            ER_774 : Bool;   // Störung Hubantrieb FU 2: Reserve
            ER_775 : Bool;   // Störung Hubantrieb FU 2: Reserve
            ER_776_ : Bool;   // Störung Hubantrieb FU 2: Reserve
            ER_777 : Bool;   // Störung Hubantrieb FU 2: Reserve
            ER_778 : Bool;   // Störung Hubantrieb FU 2: Reserve
            ER_779 : Bool;   // Störung Hubantrieb FU 2: Reserve
            ER_780 : Bool;   // Störung Hubantrieb FU 2: Reserve
         END_STRUCT;
         Reserve_1 : Struct
            ER_401 : Bool;   // Reserve
            ER_402 : Bool;   // Reserve
            ER_403 : Bool;   // Reserve
            ER_404 : Bool;   // Reserve
            ER_405 : Bool;   // Reserve
            ER_406 : Bool;   // Reserve
            ER_407 : Bool;   // Reserve
            ER_408 : Bool;   // Reserve
            ER_409 : Bool;   // Reserve
            ER_410 : Bool;   // Reserve
            ER_411 : Bool;   // Reserve
            ER_412 : Bool;   // Reserve
            ER_413 : Bool;   // Reserve
            ER_414 : Bool;   // Reserve
            ER_415 : Bool;   // Reserve
            ER_416 : Bool;   // Reserve
         END_STRUCT;
         Reserve_2 : Struct
            ER_417 : Bool;   // Reserve
            ER_418 : Bool;   // Reserve
            ER_419 : Bool;   // Reserve
            ER_420 : Bool;   // Reserve
            ER_421 : Bool;   // Reserve
            ER_422 : Bool;   // Reserve
            ER_423 : Bool;   // Reserve
            ER_424 : Bool;   // Reserve
            ER_425 : Bool;   // Reserve
            ER_426 : Bool;   // Reserve
            ER_427 : Bool;   // Reserve
            ER_428 : Bool;   // Reserve
            ER_429 : Bool;   // Reserve
            ER_430 : Bool;   // Reserve
            ER_431 : Bool;   // Reserve
            ER_432 : Bool;   // Reserve
         END_STRUCT;
         Reserve_3 : Struct
            ER_433 : Bool;   // Reserve
            ER_434 : Bool;   // Reserve
            ER_435 : Bool;   // Reserve
            ER_436 : Bool;   // Reserve
            ER_437 : Bool;   // Reserve
            ER_438 : Bool;   // Reserve
            ER_439 : Bool;   // Reserve
            ER_440 : Bool;   // Reserve
            ER_441 : Bool;   // Reserve
            ER_442 : Bool;   // Reserve
            ER_443 : Bool;   // Reserve
            ER_444 : Bool;   // Reserve
            ER_445 : Bool;   // Reserve
            ER_446 : Bool;   // Reserve
            ER_447 : Bool;   // Reserve
            ER_448 : Bool;   // Reserve
         END_STRUCT;
         Reserve_4 : Struct
            ER_449 : Bool;   // Reserve
            ER_450 : Bool;   // Reserve
            ER_451 : Bool;   // Reserve
            ER_452 : Bool;   // Reserve
            ER_453 : Bool;   // Reserve
            ER_454 : Bool;   // Reserve
            ER_455 : Bool;   // Reserve
            ER_456 : Bool;   // Reserve
            ER_457 : Bool;   // Reserve
            ER_458 : Bool;   // Reserve
            ER_459 : Bool;   // Reserve
            ER_460 : Bool;   // Reserve
            ER_461 : Bool;   // Reserve
            ER_462 : Bool;   // Reserve
            ER_463 : Bool;   // Reserve
            ER_464 : Bool;   // Reserve
         END_STRUCT;
         Reserve_5 : Struct
            ER_465 : Bool;   // Reserve
            ER_466 : Bool;   // Reserve
            ER_467 : Bool;   // Reserve
            ER_468 : Bool;   // Reserve
            ER_469 : Bool;   // Reserve
            ER_470 : Bool;   // Reserve
            ER_471 : Bool;   // Reserve
            ER_472 : Bool;   // Reserve
            ER_473 : Bool;   // Reserve
            ER_474 : Bool;   // Reserve
            ER_475 : Bool;   // Reserve
            ER_476 : Bool;   // Reserve
            ER_477 : Bool;   // Reserve
            ER_478 : Bool;   // Reserve
            ER_479 : Bool;   // Reserve
            ER_480 : Bool;   // Reserve
         END_STRUCT;
         Reserve_6 : Struct   // Meldungen Reserve
            ER_301 : Bool;   // Reserve
            ER_302 : Bool;   // Reserve
            ER_303 : Bool;   // Reserve
            ER_304 : Bool;   // Reserve
            ER_305 : Bool;   // Reserve
            ER_306 : Bool;   // Reserve
            ER_307 : Bool;   // Reserve
            ER_308 : Bool;   // Reserve
            ER_309 : Bool;   // Reserve
            ER_310 : Bool;   // Reserve
            ER_311 : Bool;   // Reserve
            ER_312 : Bool;   // Reserve
            ER_313 : Bool;   // Reserve
            ER_314 : Bool;   // Reserve
            ER_315 : Bool;   // Reserve
            ER_316 : Bool;   // Reserve
         END_STRUCT;
         Reserve_7 : Struct   // Meldungen Reserve
            ER_317 : Bool;   // Reserve
            ER_318 : Bool;   // Reserve
            ER_319 : Bool;   // Reserve
            ER_320 : Bool;   // Reserve
            ER_321 : Bool;   // Reserve
            ER_322 : Bool;   // Reserve
            ER_323 : Bool;   // Reserve
            ER_324 : Bool;   // Reserve
            ER_325 : Bool;   // Reserve
            ER_326 : Bool;   // Reserve
            ER_327 : Bool;   // Reserve
            ER_328 : Bool;   // Reserve
            ER_329 : Bool;   // Reserve
            ER_330 : Bool;   // Reserve
            ER_331 : Bool;   // Reserve
            ER_332 : Bool;   // Reserve
         END_STRUCT;
         Reserve_8 : Struct   // FU Reserve
            ER_333 : Bool;   // Störung Reserve FU 1: Überstrom
            ER_334 : Bool;   // Störung Reserve FU 1: Zwischenkreisspannung Überspannung
            ER_335 : Bool;   // Störung Reserve FU 1: Zwischenkreisspannung Unterspannung
            ER_336 : Bool;   // Störung Reserve FU 1: Übertemperatur Kühlkörper Wechselrichter
            ER_337 : Bool;   // Störung Reserve FU 1: Motordatenidentifikation fehlerhaft
            ER_338 : Bool;   // Störung Reserve FU 1: Erdschluss
            ER_339 : Bool;   // Störung Reserve FU 1: Reserve
            ER_340 : Bool;   // Störung Reserve FU 1: Führung durch PLC fehlt
            ER_341 : Bool;   // Störung Reserve FU 1: Reserve
            ER_342 : Bool;   // Störung Reserve FU 1: Reserve
            ER_343 : Bool;   // Störung Reserve FU 1: Reserve
            ER_344_ : Bool;   // Störung Reserve FU 1: Reserve
            ER_345 : Bool;   // Störung Reserve FU 1: Reserve
            ER_346 : Bool;   // Störung Reserve FU 1: Reserve
            ER_347 : Bool;   // Störung Reserve FU 1: Reserve
            ER_348 : Bool;   // Störung Reserve FU 1: Reserve
         END_STRUCT;
         Reserve_9 : Struct
            ER_349 : Bool;   // Reserve
            ER_350 : Bool;   // Reserve
            ER_351 : Bool;   // Reserve
            ER_352 : Bool;   // Reserve
            ER_353 : Bool;   // Reserve
            ER_354 : Bool;   // Reserve
            ER_355 : Bool;   // Reserve
            ER_356 : Bool;   // Reserve
            ER_357 : Bool;   // Reserve
            ER_358 : Bool;   // Reserve
            ER_359 : Bool;   // Reserve
            ER_360 : Bool;   // Reserve
            ER_361 : Bool;   // Reserve
            ER_362 : Bool;   // Reserve
            ER_363 : Bool;   // Reserve
            ER_364 : Bool;   // Reserve
         END_STRUCT;
         Reserve_10 : Struct   // FU Reserve
            ER_365 : Bool;   // Störung Reserve FU 2: Überstrom
            ER_366 : Bool;   // Störung Reserve FU 2: Zwischenkreisspannung Überspannung
            ER_367 : Bool;   // Störung Reserve FU 2: Zwischenkreisspannung Unterspannung
            ER_368 : Bool;   // Störung Reserve FU 2: Übertemperatur Kühlkörper Wechselrichter
            ER_369 : Bool;   // Störung Reserve FU 2: Motordatenidentifikation fehlerhaft
            ER_370 : Bool;   // Störung Reserve FU 2: Erdschluss
            ER_371 : Bool;   // Störung Reserve FU 2: Reserve
            ER_372 : Bool;   // Störung Reserve FU 2: Führung durch PLC fehlt
            ER_373 : Bool;   // Störung Reserve FU 2: Reserve
            ER_374 : Bool;   // Störung Reserve FU 2: Reserve
            ER_375 : Bool;   // Störung Reserve FU 2: Reserve
            ER_376 : Bool;   // Störung Reserve FU 2: Reserve
            ER_377 : Bool;   // Störung Reserve FU 2: Reserve
            ER_378 : Bool;   // Störung Reserve FU 2: Reserve
            ER_379 : Bool;   // Störung Reserve FU 2: Reserve
            ER_380 : Bool;   // Störung Reserve FU 2: Reserve
         END_STRUCT;
         SDC : Struct   // SDC Störungs
            ER_901 : Bool;   // Reserve
            ER_902 : Bool;   // Reserve
            ER_903 : Bool;   // Störung SDC Positionssprung
            ER_904 : Bool;   // Störung SDC keine Sektion gefunden
            ER_905 : Bool;   // Störung SDC Kommandos nicht plausibel
            ER_906 : Bool;   // Störung SDC Positionsgrenzen
            ER_907 : Bool;   // Störung SDC falsche EMS Nummer
            ER_908 : Bool;   // Störung SDC falsche Sektion Nummer
            ER_909 : Bool;   // Reserve
            ER_910 : Bool;   // Reserve
            ER_911 : Bool;   // Reserve
            ER_912 : Bool;   // Reserve
            ER_913 : Bool;   // Reserve
            ER_914 : Bool;   // Reserve
            ER_915 : Bool;   // Reserve
            ER_916 : Bool;   // Reserve
         END_STRUCT;
      END_STRUCT;
      EMS_ER_WORDs : Array[1..200] of Struct   // EMS Störung WORDs
         ER_WORD : Array[0..24] of Word;   // Störworte
      END_STRUCT;
      SDC : Struct
         ER_917 : Bool;   // Störung SDC Kommunikation mit Anlagensteuerung
         ER_918 : Bool;   // Störung SDC Safety Kommunikation mit Anlagensteuerung
         ER_919 : Bool;   // Störung SDC Reserve
         ER_920 : Bool;   // Störung SDC Reserve
         ER_921 : Bool;   // Störung SDC Reserve
         ER_922 : Bool;   // Störung SDC Reserve
         ER_923 : Bool;   // Störung SDC Reserve
         ER_924 : Bool;   // Störung SDC Reserve
         ER_925 : Bool;   // Störung SDC OB80 Zykluszeit
         ER_926 : Bool;   // Störung SDC OB82 Diagnosealarm
         ER_927 : Bool;   // Störung SDC OB83 Baugruppenwechsel
         ER_928 : Bool;   // Störung SDC OB86 Baugruppenträger ausgefallen
         ER_929 : Bool;   // Störung SDC OB121 Programmierfehler
         ER_930 : Bool;   // Störung SDC OB122 Peripherie-Zugriff
         ER_931 : Bool;   // Störung SDC Reserve
         ER_932 : Bool;   // Störung SDC Reserve
      END_STRUCT;
   END_VAR
BEGIN
END_DATA_BLOCK

DATA_BLOCK "DB_SDC_ERRORS_STAT"   // DB3724
{ S7_Optimized_Access := 'FALSE' }
VERSION : 0.1
   VAR
      HEADER : Struct   // Struktur für Datenheader // nicht verschieben
         DB_NR : Int := 3724;   // DB Nummer
         MIN_NR_FAULT_STAT : Int := 1;   // Niedrigste Fehler Nummer im Daten DB
         MAX_NR_FAULT_STAT : Int := 200;   // Höchste Fehler Nummer im Daten DB
         START_FAULT_STAT : Int := 20;   // Startadresse der Fehler Daten im Daten DB
         LAENGE_FAULT_STAT : Int := 28;   // Länge Fehler Daten
         FAULT_PRO_SEITE_HMI : Int := 10;   // Reserve
         RES12 : Int := 0;   // Reserve
         RES14 : Int := 0;   // Reserve
         RES16 : Int := 0;   // Reserve
         LOAD : Bool := FALSE;   // "0" zum laden des DB auf CPU
         RESET_ARCH : Bool := FALSE;   // Archiv löschen
      END_STRUCT;
      ER_ARCHIV : Array[1..1000] of "UDT_SDC_ERROR_STAT";   // Error Archiv
      ER_AKT : Array[1..200] of Struct   // Error aktiv EMS
         ER_TRIGER : Word;   // Error auslösen Aktiv von EMS
         ER_STAT : Array[1..4] of "UDT_SDC_TS_IF_STATUS_VAL";   // Error Status Aktiv EMS
      END_STRUCT;
   END_VAR
BEGIN
   ER_ARCHIV[1].EMS_TS_STAT_VAL.EMS_ID := 0;
   ER_ARCHIV[1].EMS_TS_STAT_VAL.PROFIL := 0;
   ER_ARCHIV[1].EMS_TS_STAT_VAL.DRIVE_POS := 0;
   ER_ARCHIV[1].EMS_TS_STAT_VAL.HOIST_POS := 0;
   ER_ARCHIV[1].EMS_TS_STAT_VAL.ERROR := 0;
   ER_ARCHIV[1].EMS_TS_STAT_VAL.DRIVE_POS_PERC := 0;
   ER_ARCHIV[1].EMS_TS_STAT_VAL.SEK := 0;
   ER_ARCHIV[1].ER._901_ER_SUM := FALSE;
   ER_ARCHIV[1].ER._902_ER_SUM_SDC := FALSE;
   ER_ARCHIV[1].ER._903_ER_BC_JUMP := FALSE;
   ER_ARCHIV[1].ER._904_ER_NO_SEK := FALSE;
   ER_ARCHIV[1].ER._905_ER_COMMAND := FALSE;
   ER_ARCHIV[1].ER._906_ER_BC_LIM := FALSE;
   ER_ARCHIV[1].ER._907_ER_EMS_ID := FALSE;
   ER_ARCHIV[1].ER._908_ER_SEK_NR := FALSE;
   ER_ARCHIV[1].ER._909_ER_LIFE := FALSE;
   ER_ARCHIV[1].ER._910_ER_BUS := FALSE;
   ER_ARCHIV[1].ER._911 := FALSE;
   ER_ARCHIV[1].ER._912 := FALSE;
   ER_ARCHIV[1].ER._913 := FALSE;
   ER_ARCHIV[1].ER._914 := FALSE;
   ER_ARCHIV[1].ER._915 := FALSE;
   ER_ARCHIV[1].ER._916 := FALSE;
   ER_ARCHIV[1].Spare := 0;
   ER_ARCHIV[1].ER_DATE := DT#1990-01-01-00:00:00;
   ER_ARCHIV[2].EMS_TS_STAT_VAL.EMS_ID := 0;
   ER_ARCHIV[2].EMS_TS_STAT_VAL.PROFIL := 0;
   ER_ARCHIV[2].EMS_TS_STAT_VAL.DRIVE_POS := 0;
   ER_ARCHIV[2].EMS_TS_STAT_VAL.HOIST_POS := 0;
   ER_ARCHIV[2].EMS_TS_STAT_VAL.ERROR := 0;
   ER_ARCHIV[2].EMS_TS_STAT_VAL.DRIVE_POS_PERC := 0;
   ER_ARCHIV[2].EMS_TS_STAT_VAL.SEK := 0;
   ER_ARCHIV[2].ER._901_ER_SUM := FALSE;
   ER_ARCHIV[2].ER._902_ER_SUM_SDC := FALSE;
   ER_ARCHIV[2].ER._903_ER_BC_JUMP := FALSE;
   ER_ARCHIV[2].ER._904_ER_NO_SEK := FALSE;
   ER_ARCHIV[2].ER._905_ER_COMMAND := FALSE;
   ER_ARCHIV[2].ER._906_ER_BC_LIM := FALSE;
   ER_ARCHIV[2].ER._907_ER_EMS_ID := FALSE;
   ER_ARCHIV[2].ER._908_ER_SEK_NR := FALSE;
   ER_ARCHIV[2].ER._909_ER_LIFE := FALSE;
   ER_ARCHIV[2].ER._910_ER_BUS := FALSE;
   ER_ARCHIV[2].ER._911 := FALSE;
   ER_ARCHIV[2].ER._912 := FALSE;
   ER_ARCHIV[2].ER._913 := FALSE;
   ER_ARCHIV[2].ER._914 := FALSE;
   ER_ARCHIV[2].ER._915 := FALSE;
   ER_ARCHIV[2].ER._916 := FALSE;
   ER_ARCHIV[2].Spare := 0;
   ER_ARCHIV[2].ER_DATE := DT#1990-01-01-00:00:00;
   ER_ARCHIV[3].EMS_TS_STAT_VAL.EMS_ID := 0;
   ER_ARCHIV[3].EMS_TS_STAT_VAL.PROFIL := 0;
   ER_ARCHIV[3].EMS_TS_STAT_VAL.DRIVE_POS := 0;
   ER_ARCHIV[3].EMS_TS_STAT_VAL.HOIST_POS := 0;
   ER_ARCHIV[3].EMS_TS_STAT_VAL.ERROR := 0;
   ER_ARCHIV[3].EMS_TS_STAT_VAL.DRIVE_POS_PERC := 0;
   ER_ARCHIV[3].EMS_TS_STAT_VAL.SEK := 0;
   ER_ARCHIV[3].ER._901_ER_SUM := FALSE;
   ER_ARCHIV[3].ER._902_ER_SUM_SDC := FALSE;
   ER_ARCHIV[3].ER._903_ER_BC_JUMP := FALSE;
   ER_ARCHIV[3].ER._904_ER_NO_SEK := FALSE;
   ER_ARCHIV[3].ER._905_ER_COMMAND := FALSE;
   ER_ARCHIV[3].ER._906_ER_BC_LIM := FALSE;
   ER_ARCHIV[3].ER._907_ER_EMS_ID := FALSE;
   ER_ARCHIV[3].ER._908_ER_SEK_NR := FALSE;
   ER_ARCHIV[3].ER._909_ER_LIFE := FALSE;
   ER_ARCHIV[3].ER._910_ER_BUS := FALSE;
   ER_ARCHIV[3].ER._911 := FALSE;
   ER_ARCHIV[3].ER._912 := FALSE;
   ER_ARCHIV[3].ER._913 := FALSE;
   ER_ARCHIV[3].ER._914 := FALSE;
   ER_ARCHIV[3].ER._915 := FALSE;
   ER_ARCHIV[3].ER._916 := FALSE;
   ER_ARCHIV[3].Spare := 0;
   ER_ARCHIV[3].ER_DATE := DT#1990-01-01-00:00:00;
   ER_ARCHIV[4].EMS_TS_STAT_VAL.EMS_ID := 0;
   ER_ARCHIV[4].EMS_TS_STAT_VAL.PROFIL := 0;
   ER_ARCHIV[4].EMS_TS_STAT_VAL.DRIVE_POS := 0;
   ER_ARCHIV[4].EMS_TS_STAT_VAL.HOIST_POS := 0;
   ER_ARCHIV[4].EMS_TS_STAT_VAL.ERROR := 0;
   ER_ARCHIV[4].EMS_TS_STAT_VAL.DRIVE_POS_PERC := 0;
   ER_ARCHIV[4].EMS_TS_STAT_VAL.SEK := 0;
   ER_ARCHIV[4].ER._901_ER_SUM := FALSE;
   ER_ARCHIV[4].ER._902_ER_SUM_SDC := FALSE;
   ER_ARCHIV[4].ER._903_ER_BC_JUMP := FALSE;
   ER_ARCHIV[4].ER._904_ER_NO_SEK := FALSE;
   ER_ARCHIV[4].ER._905_ER_COMMAND := FALSE;
   ER_ARCHIV[4].ER._906_ER_BC_LIM := FALSE;
   ER_ARCHIV[4].ER._907_ER_EMS_ID := FALSE;
   ER_ARCHIV[4].ER._908_ER_SEK_NR := FALSE;
   ER_ARCHIV[4].ER._909_ER_LIFE := FALSE;
   ER_ARCHIV[4].ER._910_ER_BUS := FALSE;
   ER_ARCHIV[4].ER._911 := FALSE;
   ER_ARCHIV[4].ER._912 := FALSE;
   ER_ARCHIV[4].ER._913 := FALSE;
   ER_ARCHIV[4].ER._914 := FALSE;
   ER_ARCHIV[4].ER._915 := FALSE;
   ER_ARCHIV[4].ER._916 := FALSE;
   ER_ARCHIV[4].Spare := 0;
   ER_ARCHIV[4].ER_DATE := DT#1990-01-01-00:00:00;
   ER_ARCHIV[5].EMS_TS_STAT_VAL.EMS_ID := 0;
   ER_ARCHIV[5].EMS_TS_STAT_VAL.PROFIL := 0;
   ER_ARCHIV[5].EMS_TS_STAT_VAL.DRIVE_POS := 0;
   ER_ARCHIV[5].EMS_TS_STAT_VAL.HOIST_POS := 0;
   ER_ARCHIV[5].EMS_TS_STAT_VAL.ERROR := 0;
   ER_ARCHIV[5].EMS_TS_STAT_VAL.DRIVE_POS_PERC := 0;
   ER_ARCHIV[5].EMS_TS_STAT_VAL.SEK := 0;
   ER_ARCHIV[5].ER._901_ER_SUM := FALSE;
   ER_ARCHIV[5].ER._902_ER_SUM_SDC := FALSE;
   ER_ARCHIV[5].ER._903_ER_BC_JUMP := FALSE;
   ER_ARCHIV[5].ER._904_ER_NO_SEK := FALSE;
   ER_ARCHIV[5].ER._905_ER_COMMAND := FALSE;
   ER_ARCHIV[5].ER._906_ER_BC_LIM := FALSE;
   ER_ARCHIV[5].ER._907_ER_EMS_ID := FALSE;
   ER_ARCHIV[5].ER._908_ER_SEK_NR := FALSE;
   ER_ARCHIV[5].ER._909_ER_LIFE := FALSE;
   ER_ARCHIV[5].ER._910_ER_BUS := FALSE;
   ER_ARCHIV[5].ER._911 := FALSE;
   ER_ARCHIV[5].ER._912 := FALSE;
   ER_ARCHIV[5].ER._913 := FALSE;
   ER_ARCHIV[5].ER._914 := FALSE;
   ER_ARCHIV[5].ER._915 := FALSE;
   ER_ARCHIV[5].ER._916 := FALSE;
   ER_ARCHIV[5].Spare := 0;
   ER_ARCHIV[5].ER_DATE := DT#1990-01-01-00:00:00;
   ER_ARCHIV[6].EMS_TS_STAT_VAL.EMS_ID := 0;
   ER_ARCHIV[6].EMS_TS_STAT_VAL.PROFIL := 0;
   ER_ARCHIV[6].EMS_TS_STAT_VAL.DRIVE_POS := 0;
   ER_ARCHIV[6].EMS_TS_STAT_VAL.HOIST_POS := 0;
   ER_ARCHIV[6].EMS_TS_STAT_VAL.ERROR := 0;
   ER_ARCHIV[6].EMS_TS_STAT_VAL.DRIVE_POS_PERC := 0;
   ER_ARCHIV[6].EMS_TS_STAT_VAL.SEK := 0;
   ER_ARCHIV[6].ER._901_ER_SUM := FALSE;
   ER_ARCHIV[6].ER._902_ER_SUM_SDC := FALSE;
   ER_ARCHIV[6].ER._903_ER_BC_JUMP := FALSE;
   ER_ARCHIV[6].ER._904_ER_NO_SEK := FALSE;
   ER_ARCHIV[6].ER._905_ER_COMMAND := FALSE;
   ER_ARCHIV[6].ER._906_ER_BC_LIM := FALSE;
   ER_ARCHIV[6].ER._907_ER_EMS_ID := FALSE;
   ER_ARCHIV[6].ER._908_ER_SEK_NR := FALSE;
   ER_ARCHIV[6].ER._909_ER_LIFE := FALSE;
   ER_ARCHIV[6].ER._910_ER_BUS := FALSE;
   ER_ARCHIV[6].ER._911 := FALSE;
   ER_ARCHIV[6].ER._912 := FALSE;
   ER_ARCHIV[6].ER._913 := FALSE;
   ER_ARCHIV[6].ER._914 := FALSE;
   ER_ARCHIV[6].ER._915 := FALSE;
   ER_ARCHIV[6].ER._916 := FALSE;
   ER_ARCHIV[6].Spare := 0;
   ER_ARCHIV[6].ER_DATE := DT#1990-01-01-00:00:00;
   ER_ARCHIV[7].EMS_TS_STAT_VAL.EMS_ID := 0;
   ER_ARCHIV[7].EMS_TS_STAT_VAL.PROFIL := 0;
   ER_ARCHIV[7].EMS_TS_STAT_VAL.DRIVE_POS := 0;
   ER_ARCHIV[7].EMS_TS_STAT_VAL.HOIST_POS := 0;
   ER_ARCHIV[7].EMS_TS_STAT_VAL.ERROR := 0;
   ER_ARCHIV[7].EMS_TS_STAT_VAL.DRIVE_POS_PERC := 0;
   ER_ARCHIV[7].EMS_TS_STAT_VAL.SEK := 0;
   ER_ARCHIV[7].ER._901_ER_SUM := FALSE;
   ER_ARCHIV[7].ER._902_ER_SUM_SDC := FALSE;
   ER_ARCHIV[7].ER._903_ER_BC_JUMP := FALSE;
   ER_ARCHIV[7].ER._904_ER_NO_SEK := FALSE;
   ER_ARCHIV[7].ER._905_ER_COMMAND := FALSE;
   ER_ARCHIV[7].ER._906_ER_BC_LIM := FALSE;
   ER_ARCHIV[7].ER._907_ER_EMS_ID := FALSE;
   ER_ARCHIV[7].ER._908_ER_SEK_NR := FALSE;
   ER_ARCHIV[7].ER._909_ER_LIFE := FALSE;
   ER_ARCHIV[7].ER._910_ER_BUS := FALSE;
   ER_ARCHIV[7].ER._911 := FALSE;
   ER_ARCHIV[7].ER._912 := FALSE;
   ER_ARCHIV[7].ER._913 := FALSE;
   ER_ARCHIV[7].ER._914 := FALSE;
   ER_ARCHIV[7].ER._915 := FALSE;
   ER_ARCHIV[7].ER._916 := FALSE;
   ER_ARCHIV[7].Spare := 0;
   ER_ARCHIV[7].ER_DATE := DT#1990-01-01-00:00:00;
   ER_ARCHIV[8].EMS_TS_STAT_VAL.EMS_ID := 0;
   ER_ARCHIV[8].EMS_TS_STAT_VAL.PROFIL := 0;
   ER_ARCHIV[8].EMS_TS_STAT_VAL.DRIVE_POS := 0;
   ER_ARCHIV[8].EMS_TS_STAT_VAL.HOIST_POS := 0;
   ER_ARCHIV[8].EMS_TS_STAT_VAL.ERROR := 0;
   ER_ARCHIV[8].EMS_TS_STAT_VAL.DRIVE_POS_PERC := 0;
   ER_ARCHIV[8].EMS_TS_STAT_VAL.SEK := 0;
   ER_ARCHIV[8].ER._901_ER_SUM := FALSE;
   ER_ARCHIV[8].ER._902_ER_SUM_SDC := FALSE;
   ER_ARCHIV[8].ER._903_ER_BC_JUMP := FALSE;
   ER_ARCHIV[8].ER._904_ER_NO_SEK := FALSE;
   ER_ARCHIV[8].ER._905_ER_COMMAND := FALSE;
   ER_ARCHIV[8].ER._906_ER_BC_LIM := FALSE;
   ER_ARCHIV[8].ER._907_ER_EMS_ID := FALSE;
   ER_ARCHIV[8].ER._908_ER_SEK_NR := FALSE;
   ER_ARCHIV[8].ER._909_ER_LIFE := FALSE;
   ER_ARCHIV[8].ER._910_ER_BUS := FALSE;
   ER_ARCHIV[8].ER._911 := FALSE;
   ER_ARCHIV[8].ER._912 := FALSE;
   ER_ARCHIV[8].ER._913 := FALSE;
   ER_ARCHIV[8].ER._914 := FALSE;
   ER_ARCHIV[8].ER._915 := FALSE;
   ER_ARCHIV[8].ER._916 := FALSE;
   ER_ARCHIV[8].Spare := 0;
   ER_ARCHIV[8].ER_DATE := DT#1990-01-01-00:00:00;
   // 30600 more start values not shown
END_DATA_BLOCK

DATA_BLOCK "DB_SDC_EMS_SIM"   // DB3726
{ S7_Optimized_Access := 'FALSE' }
VERSION : 0.1
   VAR
      HEADER : Struct   // Struktur für Datenheader // nicht verschieben
         DB_NR : Int := 3726;   // DB Nummer
         MIN_NR_EMS : Int := 1;   // Niedrigste EMS Nummer im Daten DB
         MAX_NR_EMS : Int := 200;   // Höchste EMS Nummer im Daten DB
         START_DAT : Int := 40;   // Startadresse der EMS Daten im Daten DB
         LAENGE_EMS : Int := 40;   // Länge Eingänge pro EMS
         RES10 : Int := 0;   // Reserve
         RES12 : Int := 0;   // Reserve
         RES14 : Int := 0;   // Reserve
         RES16 : Int := 0;   // Reserve
         RES18 : Int := 0;   // Reserve
      END_STRUCT;
      PAR : Struct   // Parameter Simulation
         BARCODE_START : DInt := 1;   // min Barcodevalue
         BARCODE_ENDE : DInt := 500000;   // max Barcodevalue
         HUB_START : Int := 0;   // min Hoistvalue
         HUB_ENDE : Int := 4010;   // max Hoistvalue
         LEAP_AKT : Array[1..20] of Bool;   // Leap Aktiv
         LEAP_HIGH_LOW : Array[1..20] of Bool;   // Leap Aktiv
         ON : Bool := TRUE;   // Simulation ON "1"
         RES18 : Int := 0;   // Reserve
      END_STRUCT;
      EMS : Array[1..200] of "UDT_EMS_IF_Q";   // EMS Simulation Eingänge
      EMS_TEMP : "UDT_EMS_IF_Q";
   END_VAR
BEGIN
   PAR.LEAP_AKT[1] := TRUE;
   PAR.LEAP_AKT[2] := TRUE;
   PAR.LEAP_AKT[3] := TRUE;
   PAR.LEAP_HIGH_LOW[1] := TRUE;
   PAR.LEAP_HIGH_LOW[2] := FALSE;
   PAR.LEAP_HIGH_LOW[3] := TRUE;
   PAR.LEAP_AKT[4] := FALSE;
   PAR.LEAP_AKT[5] := FALSE;
   PAR.LEAP_AKT[6] := FALSE;
   PAR.LEAP_AKT[7] := FALSE;
   PAR.LEAP_AKT[8] := FALSE;
   PAR.LEAP_AKT[9] := FALSE;
   PAR.LEAP_AKT[10] := FALSE;
   PAR.LEAP_AKT[11] := FALSE;
   PAR.LEAP_AKT[12] := FALSE;
   PAR.LEAP_AKT[13] := FALSE;
   PAR.LEAP_AKT[14] := FALSE;
   PAR.LEAP_AKT[15] := FALSE;
   PAR.LEAP_AKT[16] := FALSE;
   PAR.LEAP_AKT[17] := FALSE;
   PAR.LEAP_AKT[18] := FALSE;
   PAR.LEAP_AKT[19] := FALSE;
   PAR.LEAP_AKT[20] := FALSE;
   PAR.LEAP_HIGH_LOW[4] := FALSE;
   PAR.LEAP_HIGH_LOW[5] := FALSE;
   PAR.LEAP_HIGH_LOW[6] := FALSE;
   PAR.LEAP_HIGH_LOW[7] := FALSE;
   PAR.LEAP_HIGH_LOW[8] := FALSE;
   PAR.LEAP_HIGH_LOW[9] := FALSE;
   PAR.LEAP_HIGH_LOW[10] := FALSE;
   PAR.LEAP_HIGH_LOW[11] := FALSE;
   PAR.LEAP_HIGH_LOW[12] := FALSE;
   PAR.LEAP_HIGH_LOW[13] := FALSE;
   PAR.LEAP_HIGH_LOW[14] := FALSE;
   PAR.LEAP_HIGH_LOW[15] := FALSE;
   PAR.LEAP_HIGH_LOW[16] := FALSE;
   PAR.LEAP_HIGH_LOW[17] := FALSE;
   PAR.LEAP_HIGH_LOW[18] := FALSE;
   PAR.LEAP_HIGH_LOW[19] := FALSE;
   PAR.LEAP_HIGH_LOW[20] := FALSE;
   EMS[1].STAT.LIFE_BIT := TRUE;
   EMS[1].STAT.ER_SUM := FALSE;
   EMS[1].STAT.IR_MAN := FALSE;
   EMS[1].STAT.ER_RESET := FALSE;
   EMS[1].STAT.HOIST_CLEAR := FALSE;
   EMS[1].STAT.POS_START_X := FALSE;
   EMS[1].STAT.ALWAYS_ONE := TRUE;
   EMS[1].STAT.H_DISABLED := FALSE;
   EMS[1].STAT.D_FWD := TRUE;
   EMS[1].STAT.D_RWD := FALSE;
   EMS[1].STAT.bit12 := FALSE;
   EMS[1].STAT.D_IN_POS := FALSE;
   EMS[1].STAT.H_UP := FALSE;
   EMS[1].STAT.H_DOWN := FALSE;
   EMS[1].STAT.H_IN_POS := TRUE;
   EMS[1].STAT.H_IN_TOPPOS := FALSE;
   EMS[1].STAT.bit2_0 := FALSE;
   EMS[1].STAT.bit2_1 := FALSE;
   EMS[1].STAT.bit2_2 := FALSE;
   EMS[1].STAT.bit2_3 := FALSE;
   EMS[1].STAT.IN_BOTPOS := FALSE;
   EMS[1].STAT.bit2_5 := FALSE;
   EMS[1].STAT.bit2_6 := FALSE;
   EMS[1].STAT.bit2_7 := FALSE;
   EMS[1].STAT.MESS_POS := FALSE;
   EMS[1].STAT.bit3_2 := FALSE;
   EMS[1].STAT.bit3_3 := FALSE;
   EMS[1].STAT.bit3_4 := FALSE;
   EMS[1].STAT.bit3_5 := FALSE;
   EMS[1].STAT.bit3_6 := FALSE;
   EMS[1].STAT.DATA_TRANS := FALSE;
   EMS[1].ERROR := 0;
   EMS[1].D_POS := 22899;
   EMS[1].H_POS := 603;
   EMS[1].ER_WORD_No := 1;
   EMS[1].ER_WORD := 16#0000;
   EMS[1].FB_DBNo := 0;
   EMS[1].FB_DBBNo := 0;
   EMS[2].STAT.LIFE_BIT := TRUE;
   EMS[2].STAT.ER_SUM := FALSE;
   EMS[2].STAT.IR_MAN := FALSE;
   EMS[2].STAT.ER_RESET := FALSE;
   EMS[2].STAT.HOIST_CLEAR := FALSE;
   EMS[2].STAT.POS_START_X := FALSE;
   EMS[2].STAT.ALWAYS_ONE := TRUE;
   EMS[2].STAT.H_DISABLED := FALSE;
   EMS[2].STAT.D_FWD := TRUE;
   EMS[2].STAT.D_RWD := FALSE;
   EMS[2].STAT.bit12 := FALSE;
   EMS[2].STAT.D_IN_POS := FALSE;
   EMS[2].STAT.H_UP := FALSE;
   EMS[2].STAT.H_DOWN := FALSE;
   EMS[2].STAT.H_IN_POS := FALSE;
   EMS[2].STAT.H_IN_TOPPOS := TRUE;
   EMS[2].STAT.bit2_0 := FALSE;
   EMS[2].STAT.bit2_1 := FALSE;
   EMS[2].STAT.bit2_2 := FALSE;
   EMS[2].STAT.bit2_3 := FALSE;
   EMS[2].STAT.IN_BOTPOS := FALSE;
   EMS[2].STAT.bit2_5 := FALSE;
   EMS[2].STAT.bit2_6 := FALSE;
   EMS[2].STAT.bit2_7 := FALSE;
   EMS[2].STAT.MESS_POS := FALSE;
   EMS[2].STAT.bit3_2 := FALSE;
   EMS[2].STAT.bit3_3 := FALSE;
   EMS[2].STAT.bit3_4 := FALSE;
   EMS[2].STAT.bit3_5 := FALSE;
   EMS[2].STAT.bit3_6 := FALSE;
   EMS[2].STAT.DATA_TRANS := FALSE;
   EMS[2].ERROR := 0;
   EMS[2].D_POS := 10522;
   EMS[2].H_POS := 4010;
   EMS[2].ER_WORD_No := 1;
   EMS[2].ER_WORD := 16#0000;
   EMS[2].FB_DBNo := 0;
   EMS[2].FB_DBBNo := 0;
   EMS[3].STAT.LIFE_BIT := TRUE;
   EMS[3].STAT.ER_SUM := FALSE;
   EMS[3].STAT.IR_MAN := FALSE;
   EMS[3].STAT.ER_RESET := FALSE;
   EMS[3].STAT.HOIST_CLEAR := FALSE;
   EMS[3].STAT.POS_START_X := FALSE;
   EMS[3].STAT.ALWAYS_ONE := TRUE;
   EMS[3].STAT.H_DISABLED := FALSE;
   EMS[3].STAT.D_FWD := TRUE;
   EMS[3].STAT.D_RWD := FALSE;
   EMS[3].STAT.bit12 := FALSE;
   EMS[3].STAT.D_IN_POS := FALSE;
   EMS[3].STAT.H_UP := FALSE;
   EMS[3].STAT.H_DOWN := FALSE;
   EMS[3].STAT.H_IN_POS := FALSE;
   EMS[3].STAT.H_IN_TOPPOS := TRUE;
   EMS[3].STAT.bit2_0 := FALSE;
   EMS[3].STAT.bit2_1 := FALSE;
   EMS[3].STAT.bit2_2 := FALSE;
   EMS[3].STAT.bit2_3 := FALSE;
   EMS[3].STAT.IN_BOTPOS := FALSE;
   EMS[3].STAT.bit2_5 := FALSE;
   EMS[3].STAT.bit2_6 := FALSE;
   EMS[3].STAT.bit2_7 := FALSE;
   EMS[3].STAT.MESS_POS := FALSE;
   EMS[3].STAT.bit3_2 := FALSE;
   EMS[3].STAT.bit3_3 := FALSE;
   EMS[3].STAT.bit3_4 := FALSE;
   EMS[3].STAT.bit3_5 := FALSE;
   EMS[3].STAT.bit3_6 := FALSE;
   EMS[3].STAT.DATA_TRANS := FALSE;
   EMS[3].ERROR := 0;
   EMS[3].D_POS := 96650;
   EMS[3].H_POS := 4010;
   EMS[3].ER_WORD_No := 1;
   EMS[3].ER_WORD := 16#0000;
   EMS[3].FB_DBNo := 0;
   EMS[3].FB_DBBNo := 0;
   EMS[4].STAT.LIFE_BIT := FALSE;
   EMS[4].STAT.ER_SUM := FALSE;
   EMS[4].STAT.IR_MAN := FALSE;
   EMS[4].STAT.ER_RESET := FALSE;
   EMS[4].STAT.HOIST_CLEAR := FALSE;
   EMS[4].STAT.POS_START_X := FALSE;
   EMS[4].STAT.ALWAYS_ONE := FALSE;
   EMS[4].STAT.H_DISABLED := FALSE;
   EMS[4].STAT.D_FWD := FALSE;
   EMS[4].STAT.D_RWD := FALSE;
   EMS[4].STAT.bit12 := FALSE;
   EMS[4].STAT.D_IN_POS := FALSE;
   EMS[4].STAT.H_UP := FALSE;
   EMS[4].STAT.H_DOWN := FALSE;
   EMS[4].STAT.H_IN_POS := FALSE;
   EMS[4].STAT.H_IN_TOPPOS := FALSE;
   EMS[4].STAT.bit2_0 := FALSE;
   EMS[4].STAT.bit2_1 := FALSE;
   EMS[4].STAT.bit2_2 := FALSE;
   EMS[4].STAT.bit2_3 := FALSE;
   EMS[4].STAT.IN_BOTPOS := FALSE;
   EMS[4].STAT.bit2_5 := FALSE;
   EMS[4].STAT.bit2_6 := FALSE;
   EMS[4].STAT.bit2_7 := FALSE;
   EMS[4].STAT.MESS_POS := FALSE;
   EMS[4].STAT.bit3_2 := FALSE;
   EMS[4].STAT.bit3_3 := FALSE;
   EMS[4].STAT.bit3_4 := FALSE;
   EMS[4].STAT.bit3_5 := FALSE;
   EMS[4].STAT.bit3_6 := FALSE;
   EMS[4].STAT.DATA_TRANS := FALSE;
   EMS[4].ERROR := 0;
   EMS[4].D_POS := 0;
   EMS[4].H_POS := 0;
   EMS[4].ER_WORD_No := 0;
   EMS[4].ER_WORD := 16#0000;
   EMS[4].FB_DBNo := 0;
   EMS[4].FB_DBBNo := 0;
   EMS[5].STAT.LIFE_BIT := FALSE;
   EMS[5].STAT.ER_SUM := FALSE;
   EMS[5].STAT.IR_MAN := FALSE;
   EMS[5].STAT.ER_RESET := FALSE;
   EMS[5].STAT.HOIST_CLEAR := FALSE;
   EMS[5].STAT.POS_START_X := FALSE;
   EMS[5].STAT.ALWAYS_ONE := FALSE;
   EMS[5].STAT.H_DISABLED := FALSE;
   // 15719 more start values not shown
END_DATA_BLOCK

DATA_BLOCK "DB_SDC_EMS_TA"   // DB3728
{ S7_Optimized_Access := 'FALSE' }
VERSION : 0.1
   VAR
      HEADER : Struct
         DB_NR : Int := 3728;
         MIN_NR_EMS : Int := 1;
         MAX_NR_EMS : Int := 200;
         START_EMS : Int := 20;
         LAENGE_TA_DATA : Int := 6;
         ANZ_TA : Int := 3;
         Res120 : Int;
         Res140 : Int;
         Res160 : Int;
         Load : Bool := TRUE;
      END_STRUCT;
      EMS : Array[1..200] of Struct
         TA : Array[1..3] of "UDT_EMS_TA";
      END_STRUCT;
   END_VAR
BEGIN
END_DATA_BLOCK

DATA_BLOCK "DB_SDC_BARCODE_INSERTS"   // DB3734
{ S7_Optimized_Access := 'FALSE' }
VERSION : 0.1
   VAR
      HYST : Int := 100;   // Hysterese für Positionswerte
      INSERTS : Int := 2;   // Positioning Leaps
      INSERT : Array[1..20] of Struct   // LEAPs
         COURSELOW : DInt;   // lower position value Course Barocdevalue befor Insert
         COURSEHIGH : DInt;   // höhere Positionswert Course Barocde Wert nach Insert
         INSERTLOW : DInt;   // lower position value Barocdevalue Insert low
         INSERTHIGH : DInt;   // höhere Positionswert Barocde Wert liegt Hoch
         OFFSET : DInt;   // absoluten Offset zu Beginn der Einfügen -> zusätzlich von allen Einsätzen unter
      END_STRUCT;
      ABS_DIST_COURSE : DInt := 304270;   // abslolute Entfernung
   END_VAR
BEGIN
   INSERT[2].COURSELOW := 254280;
   INSERT[1].COURSEHIGH := 5800;
   INSERT[2].COURSEHIGH := 256410;
   INSERT[2].INSERTLOW := 0;
   INSERT[2].INSERTHIGH := 0;
   INSERT[1].OFFSET := -5800;
   INSERT[2].OFFSET := -7930;
   INSERT[1].COURSELOW := 0;
   INSERT[1].INSERTLOW := 0;
   INSERT[1].INSERTHIGH := 0;
   INSERT[3].COURSELOW := 0;
   INSERT[3].COURSEHIGH := 0;
   INSERT[3].INSERTLOW := 0;
   INSERT[3].INSERTHIGH := 0;
   INSERT[3].OFFSET := -1000;
   INSERT[4].COURSELOW := 0;
   INSERT[4].COURSEHIGH := 0;
   INSERT[4].INSERTLOW := 0;
   INSERT[4].INSERTHIGH := 0;
   INSERT[4].OFFSET := -1000;
   INSERT[5].COURSELOW := 0;
   INSERT[5].COURSEHIGH := 0;
   INSERT[5].INSERTLOW := 0;
   INSERT[5].INSERTHIGH := 0;
   INSERT[5].OFFSET := -1000;
   INSERT[6].COURSELOW := 0;
   INSERT[6].COURSEHIGH := 0;
   INSERT[6].INSERTLOW := 0;
   INSERT[6].INSERTHIGH := 0;
   INSERT[6].OFFSET := -1000;
   INSERT[7].COURSELOW := 0;
   INSERT[7].COURSEHIGH := 0;
   INSERT[7].INSERTLOW := 0;
   INSERT[7].INSERTHIGH := 0;
   INSERT[7].OFFSET := -1000;
   INSERT[8].COURSELOW := 0;
   INSERT[8].COURSEHIGH := 0;
   INSERT[8].INSERTLOW := 0;
   INSERT[8].INSERTHIGH := 0;
   INSERT[8].OFFSET := -1000;
   INSERT[9].COURSELOW := 0;
   INSERT[9].COURSEHIGH := 0;
   INSERT[9].INSERTLOW := 0;
   INSERT[9].INSERTHIGH := 0;
   INSERT[9].OFFSET := -1000;
   INSERT[10].COURSELOW := 0;
   INSERT[10].COURSEHIGH := 0;
   INSERT[10].INSERTLOW := 0;
   INSERT[10].INSERTHIGH := 0;
   INSERT[10].OFFSET := -1000;
   INSERT[11].COURSELOW := 0;
   INSERT[11].COURSEHIGH := 0;
   INSERT[11].INSERTLOW := 0;
   INSERT[11].INSERTHIGH := 0;
   INSERT[11].OFFSET := 0;
   INSERT[12].COURSELOW := 0;
   INSERT[12].COURSEHIGH := 0;
   INSERT[12].INSERTLOW := 0;
   INSERT[12].INSERTHIGH := 0;
   INSERT[12].OFFSET := 0;
   INSERT[13].COURSELOW := 0;
   INSERT[13].COURSEHIGH := 0;
   INSERT[13].INSERTLOW := 0;
   INSERT[13].INSERTHIGH := 0;
   INSERT[13].OFFSET := 0;
   INSERT[14].COURSELOW := 0;
   INSERT[14].COURSEHIGH := 0;
   INSERT[14].INSERTLOW := 0;
   INSERT[14].INSERTHIGH := 0;
   INSERT[14].OFFSET := 0;
   INSERT[15].COURSELOW := 0;
   INSERT[15].COURSEHIGH := 0;
   INSERT[15].INSERTLOW := 0;
   INSERT[15].INSERTHIGH := 0;
   INSERT[15].OFFSET := 0;
   INSERT[16].COURSELOW := 0;
   INSERT[16].COURSEHIGH := 0;
   INSERT[16].INSERTLOW := 0;
   INSERT[16].INSERTHIGH := 0;
   INSERT[16].OFFSET := 0;
   INSERT[17].COURSELOW := 0;
   INSERT[17].COURSEHIGH := 0;
   INSERT[17].INSERTLOW := 0;
   INSERT[17].INSERTHIGH := 0;
   INSERT[17].OFFSET := 0;
   INSERT[18].COURSELOW := 0;
   INSERT[18].COURSEHIGH := 0;
   INSERT[18].INSERTLOW := 0;
   INSERT[18].INSERTHIGH := 0;
   INSERT[18].OFFSET := 0;
   INSERT[19].COURSELOW := 0;
   INSERT[19].COURSEHIGH := 0;
   INSERT[19].INSERTLOW := 0;
   INSERT[19].INSERTHIGH := 0;
   INSERT[19].OFFSET := 0;
   INSERT[20].COURSELOW := 0;
   INSERT[20].COURSEHIGH := 0;
   INSERT[20].INSERTLOW := 0;
   INSERT[20].INSERTHIGH := 0;
   INSERT[20].OFFSET := 0;
END_DATA_BLOCK

